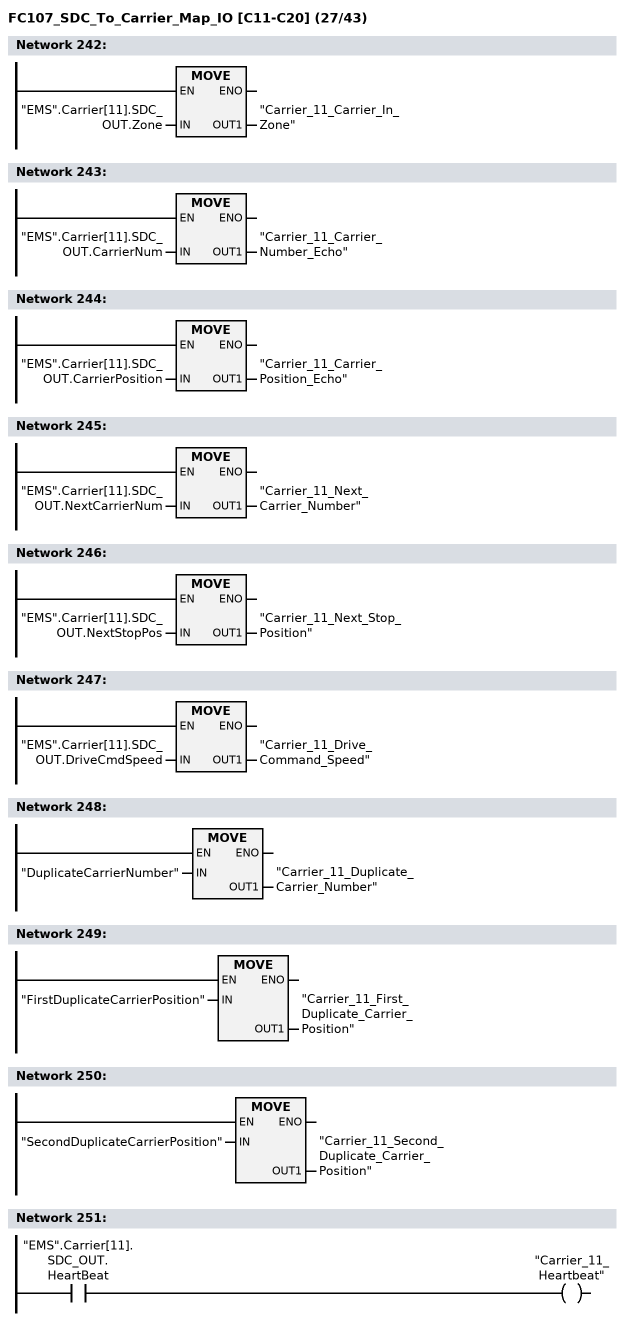
   RUNG wire#powerrail
      Move(in := "EMS".Carrier[11].SDC_OUT.Zone, out1 => "Carrier_11_Carrier_In_Zone")
   END_RUNG
   // the same network as SCL:
   "Carrier_11_Carrier_In_Zone" := "EMS".Carrier[11].SDC_OUT.Zone;
END_REGION

REGION Network 243
   RUNG wire#powerrail
      Move(in := "EMS".Carrier[11].SDC_OUT.CarrierNum, out1 => "Carrier_11_Carrier_Number_Echo")
   END_RUNG
   // the same network as SCL:
   "Carrier_11_Carrier_Number_Echo" := "EMS".Carrier[11].SDC_OUT.CarrierNum;
END_REGION

REGION Network 244
   RUNG wire#powerrail
      Move(in := "EMS".Carrier[11].SDC_OUT.CarrierPosition, out1 => "Carrier_11_Carrier_Position_Echo")
   END_RUNG
   // the same network as SCL:
   "Carrier_11_Carrier_Position_Echo" := "EMS".Carrier[11].SDC_OUT.CarrierPosition;
END_REGION

REGION Network 245
   RUNG wire#powerrail
      Move(in := "EMS".Carrier[11].SDC_OUT.NextCarrierNum, out1 => "Carrier_11_Next_Carrier_Number")
   END_RUNG
   // the same network as SCL:
   "Carrier_11_Next_Carrier_Number" := "EMS".Carrier[11].SDC_OUT.NextCarrierNum;
END_REGION

REGION Network 246
   RUNG wire#powerrail
      Move(in := "EMS".Carrier[11].SDC_OUT.NextStopPos, out1 => "Carrier_11_Next_Stop_Position")
   END_RUNG
   // the same network as SCL:
   "Carrier_11_Next_Stop_Position" := "EMS".Carrier[11].SDC_OUT.NextStopPos;
END_REGION

REGION Network 247
   RUNG wire#powerrail
      Move(in := "EMS".Carrier[11].SDC_OUT.DriveCmdSpeed, out1 => "Carrier_11_Drive_Command_Speed")
   END_RUNG
   // the same network as SCL:
   "Carrier_11_Drive_Command_Speed" := "EMS".Carrier[11].SDC_OUT.DriveCmdSpeed;
END_REGION

REGION Network 248
   RUNG wire#powerrail
      Move(in := "DuplicateCarrierNumber", out1 => "Carrier_11_Duplicate_Carrier_Number")
   END_RUNG
   // the same network as SCL:
   "Carrier_11_Duplicate_Carrier_Number" := "DuplicateCarrierNumber";
END_REGION

REGION Network 249
   RUNG wire#powerrail
      Move(in := "FirstDuplicateCarrierPosition", out1 => "Carrier_11_First_Duplicate_Carrier_Position")
   END_RUNG
   // the same network as SCL:
   "Carrier_11_First_Duplicate_Carrier_Position" := "FirstDuplicateCarrierPosition";
END_REGION

REGION Network 250
   RUNG wire#powerrail
      Move(in := "SecondDuplicateCarrierPosition", out1 => "Carrier_11_Second_Duplicate_Carrier_Position")
   END_RUNG
   // the same network as SCL:
   "Carrier_11_Second_Duplicate_Carrier_Position" := "SecondDuplicateCarrierPosition";
END_REGION

REGION Network 251
   RUNG wire#powerrail
      Contact( "EMS".Carrier[11].SDC_OUT.HeartBeat )
      Coil( "Carrier_11_Heartbeat" )
   END_RUNG
   // the same network as SCL:
   "Carrier_11_Heartbeat" := "EMS".Carrier[11].SDC_OUT.HeartBeat;
END_REGION

REGION Network 252
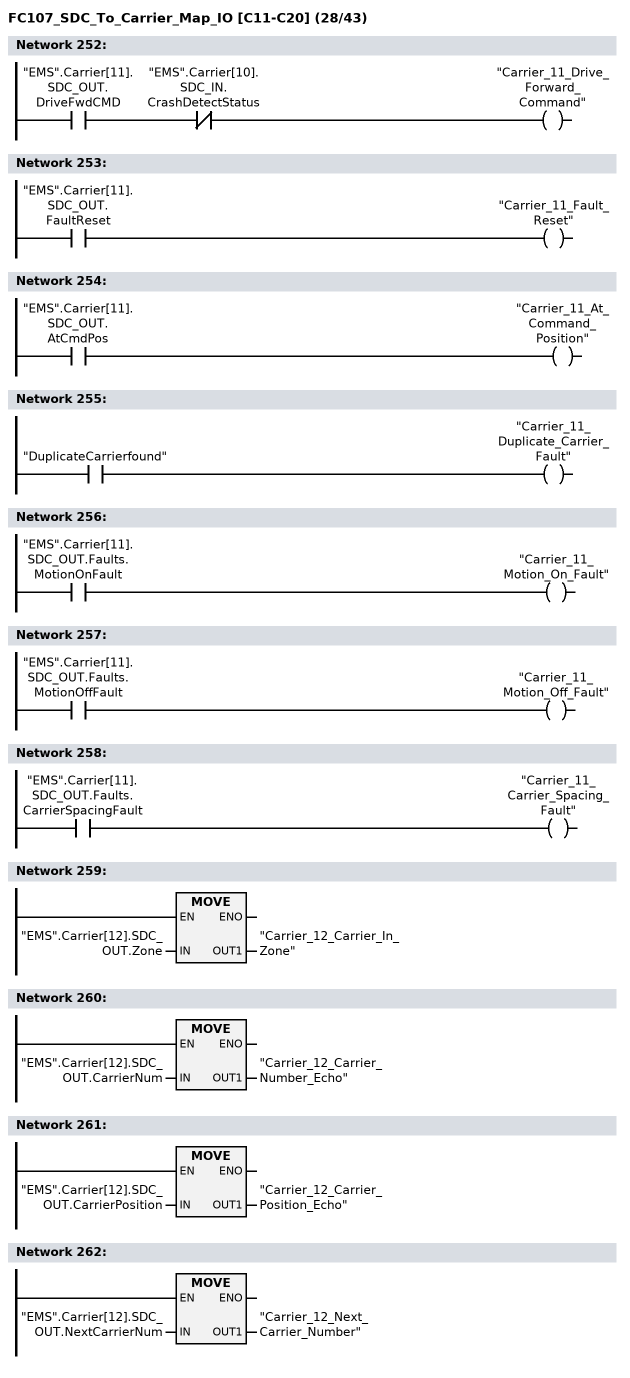
   RUNG wire#powerrail
      Contact( "EMS".Carrier[11].SDC_OUT.DriveFwdCMD )
      I_Contact( "EMS".Carrier[10].SDC_IN.CrashDetectStatus )
      Coil( "Carrier_11_Drive_Forward_Command" )
   END_RUNG
   // the same network as SCL:
   "Carrier_11_Drive_Forward_Command" := "EMS".Carrier[11].SDC_OUT.DriveFwdCMD AND NOT "EMS".Carrier[10].SDC_IN.CrashDetectStatus;
END_REGION

REGION Network 253
   RUNG wire#powerrail
      Contact( "EMS".Carrier[11].SDC_OUT.FaultReset )
      Coil( "Carrier_11_Fault_Reset" )
   END_RUNG
   // the same network as SCL:
   "Carrier_11_Fault_Reset" := "EMS".Carrier[11].SDC_OUT.FaultReset;
END_REGION

REGION Network 254
   RUNG wire#powerrail
      Contact( "EMS".Carrier[11].SDC_OUT.AtCmdPos )
      Coil( "Carrier_11_At_Command_Position" )
   END_RUNG
   // the same network as SCL:
   "Carrier_11_At_Command_Position" := "EMS".Carrier[11].SDC_OUT.AtCmdPos;
END_REGION

REGION Network 255
   RUNG wire#powerrail
      Contact( "DuplicateCarrierfound" )
      Coil( "Carrier_11_Duplicate_Carrier_Fault" )
   END_RUNG
   // the same network as SCL:
   "Carrier_11_Duplicate_Carrier_Fault" := "DuplicateCarrierfound";
END_REGION

REGION Network 256
   RUNG wire#powerrail
      Contact( "EMS".Carrier[11].SDC_OUT.Faults.MotionOnFault )
      Coil( "Carrier_11_Motion_On_Fault" )
   END_RUNG
   // the same network as SCL:
   "Carrier_11_Motion_On_Fault" := "EMS".Carrier[11].SDC_OUT.Faults.MotionOnFault;
END_REGION

REGION Network 257
   RUNG wire#powerrail
      Contact( "EMS".Carrier[11].SDC_OUT.Faults.MotionOffFault )
      Coil( "Carrier_11_Motion_Off_Fault" )
   END_RUNG
   // the same network as SCL:
   "Carrier_11_Motion_Off_Fault" := "EMS".Carrier[11].SDC_OUT.Faults.MotionOffFault;
END_REGION

REGION Network 258
   RUNG wire#powerrail
      Contact( "EMS".Carrier[11].SDC_OUT.Faults.CarrierSpacingFault )
      Coil( "Carrier_11_Carrier_Spacing_Fault" )
   END_RUNG
   // the same network as SCL:
   "Carrier_11_Carrier_Spacing_Fault" := "EMS".Carrier[11].SDC_OUT.Faults.CarrierSpacingFault;
END_REGION

REGION Network 259
   RUNG wire#powerrail
      Move(in := "EMS".Carrier[12].SDC_OUT.Zone, out1 => "Carrier_12_Carrier_In_Zone")
   END_RUNG
   // the same network as SCL:
   "Carrier_12_Carrier_In_Zone" := "EMS".Carrier[12].SDC_OUT.Zone;
END_REGION

REGION Network 260
   RUNG wire#powerrail
      Move(in := "EMS".Carrier[12].SDC_OUT.CarrierNum, out1 => "Carrier_12_Carrier_Number_Echo")
   END_RUNG
   // the same network as SCL:
   "Carrier_12_Carrier_Number_Echo" := "EMS".Carrier[12].SDC_OUT.CarrierNum;
END_REGION

REGION Network 261
   RUNG wire#powerrail
      Move(in := "EMS".Carrier[12].SDC_OUT.CarrierPosition, out1 => "Carrier_12_Carrier_Position_Echo")
   END_RUNG
   // the same network as SCL:
   "Carrier_12_Carrier_Position_Echo" := "EMS".Carrier[12].SDC_OUT.CarrierPosition;
END_REGION

REGION Network 262
   RUNG wire#powerrail
      Move(in := "EMS".Carrier[12].SDC_OUT.NextCarrierNum, out1 => "Carrier_12_Next_Carrier_Number")
   END_RUNG
   // the same network as SCL:
   "Carrier_12_Next_Carrier_Number" := "EMS".Carrier[12].SDC_OUT.NextCarrierNum;
END_REGION

REGION Network 263
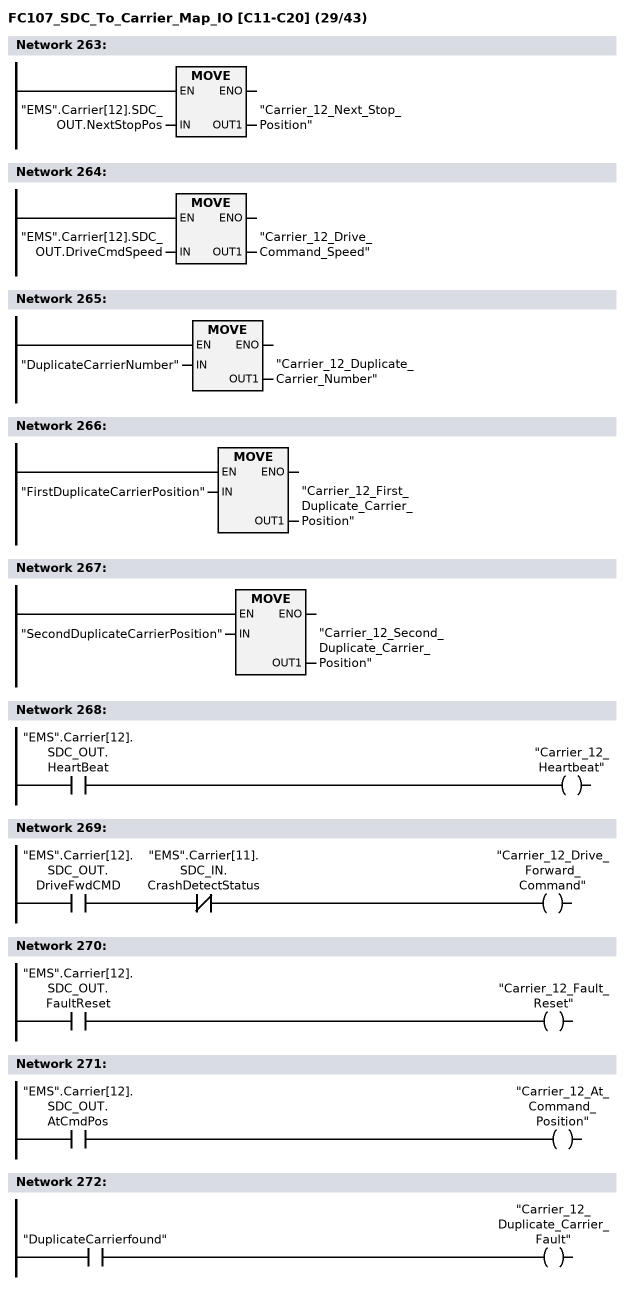
   RUNG wire#powerrail
      Move(in := "EMS".Carrier[12].SDC_OUT.NextStopPos, out1 => "Carrier_12_Next_Stop_Position")
   END_RUNG
   // the same network as SCL:
   "Carrier_12_Next_Stop_Position" := "EMS".Carrier[12].SDC_OUT.NextStopPos;
END_REGION

REGION Network 264
   RUNG wire#powerrail
      Move(in := "EMS".Carrier[12].SDC_OUT.DriveCmdSpeed, out1 => "Carrier_12_Drive_Command_Speed")
   END_RUNG
   // the same network as SCL:
   "Carrier_12_Drive_Command_Speed" := "EMS".Carrier[12].SDC_OUT.DriveCmdSpeed;
END_REGION

REGION Network 265
   RUNG wire#powerrail
      Move(in := "DuplicateCarrierNumber", out1 => "Carrier_12_Duplicate_Carrier_Number")
   END_RUNG
   // the same network as SCL:
   "Carrier_12_Duplicate_Carrier_Number" := "DuplicateCarrierNumber";
END_REGION

REGION Network 266
   RUNG wire#powerrail
      Move(in := "FirstDuplicateCarrierPosition", out1 => "Carrier_12_First_Duplicate_Carrier_Position")
   END_RUNG
   // the same network as SCL:
   "Carrier_12_First_Duplicate_Carrier_Position" := "FirstDuplicateCarrierPosition";
END_REGION

REGION Network 267
   RUNG wire#powerrail
      Move(in := "SecondDuplicateCarrierPosition", out1 => "Carrier_12_Second_Duplicate_Carrier_Position")
   END_RUNG
   // the same network as SCL:
   "Carrier_12_Second_Duplicate_Carrier_Position" := "SecondDuplicateCarrierPosition";
END_REGION

REGION Network 268
   RUNG wire#powerrail
      Contact( "EMS".Carrier[12].SDC_OUT.HeartBeat )
      Coil( "Carrier_12_Heartbeat" )
   END_RUNG
   // the same network as SCL:
   "Carrier_12_Heartbeat" := "EMS".Carrier[12].SDC_OUT.HeartBeat;
END_REGION

REGION Network 269
   RUNG wire#powerrail
      Contact( "EMS".Carrier[12].SDC_OUT.DriveFwdCMD )
      I_Contact( "EMS".Carrier[11].SDC_IN.CrashDetectStatus )
      Coil( "Carrier_12_Drive_Forward_Command" )
   END_RUNG
   // the same network as SCL:
   "Carrier_12_Drive_Forward_Command" := "EMS".Carrier[12].SDC_OUT.DriveFwdCMD AND NOT "EMS".Carrier[11].SDC_IN.CrashDetectStatus;
END_REGION

REGION Network 270
   RUNG wire#powerrail
      Contact( "EMS".Carrier[12].SDC_OUT.FaultReset )
      Coil( "Carrier_12_Fault_Reset" )
   END_RUNG
   // the same network as SCL:
   "Carrier_12_Fault_Reset" := "EMS".Carrier[12].SDC_OUT.FaultReset;
END_REGION

REGION Network 271
   RUNG wire#powerrail
      Contact( "EMS".Carrier[12].SDC_OUT.AtCmdPos )
      Coil( "Carrier_12_At_Command_Position" )
   END_RUNG
   // the same network as SCL:
   "Carrier_12_At_Command_Position" := "EMS".Carrier[12].SDC_OUT.AtCmdPos;
END_REGION

REGION Network 272
   RUNG wire#powerrail
      Contact( "DuplicateCarrierfound" )
      Coil( "Carrier_12_Duplicate_Carrier_Fault" )
   END_RUNG
   // the same network as SCL:
   "Carrier_12_Duplicate_Carrier_Fault" := "DuplicateCarrierfound";
END_REGION

REGION Network 273
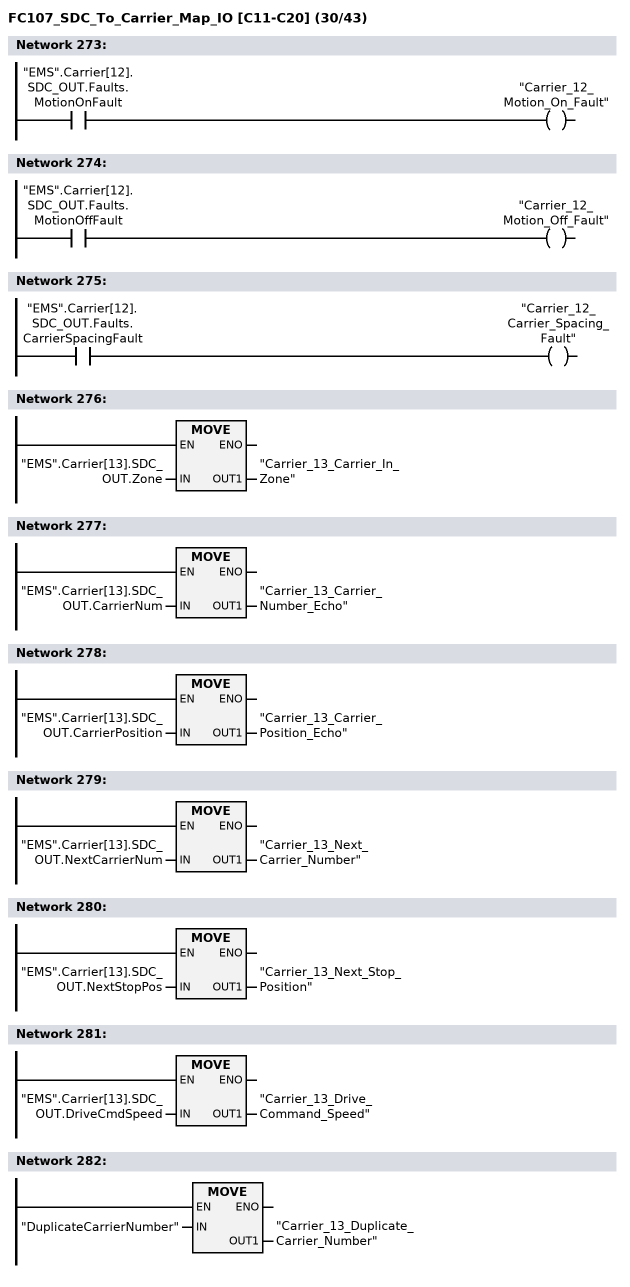
   RUNG wire#powerrail
      Contact( "EMS".Carrier[12].SDC_OUT.Faults.MotionOnFault )
      Coil( "Carrier_12_Motion_On_Fault" )
   END_RUNG
   // the same network as SCL:
   "Carrier_12_Motion_On_Fault" := "EMS".Carrier[12].SDC_OUT.Faults.MotionOnFault;
END_REGION

REGION Network 274
   RUNG wire#powerrail
      Contact( "EMS".Carrier[12].SDC_OUT.Faults.MotionOffFault )
      Coil( "Carrier_12_Motion_Off_Fault" )
   END_RUNG
   // the same network as SCL:
   "Carrier_12_Motion_Off_Fault" := "EMS".Carrier[12].SDC_OUT.Faults.MotionOffFault;
END_REGION

REGION Network 275
   RUNG wire#powerrail
      Contact( "EMS".Carrier[12].SDC_OUT.Faults.CarrierSpacingFault )
      Coil( "Carrier_12_Carrier_Spacing_Fault" )
   END_RUNG
   // the same network as SCL:
   "Carrier_12_Carrier_Spacing_Fault" := "EMS".Carrier[12].SDC_OUT.Faults.CarrierSpacingFault;
END_REGION

REGION Network 276
   RUNG wire#powerrail
      Move(in := "EMS".Carrier[13].SDC_OUT.Zone, out1 => "Carrier_13_Carrier_In_Zone")
   END_RUNG
   // the same network as SCL:
   "Carrier_13_Carrier_In_Zone" := "EMS".Carrier[13].SDC_OUT.Zone;
END_REGION

REGION Network 277
   RUNG wire#powerrail
      Move(in := "EMS".Carrier[13].SDC_OUT.CarrierNum, out1 => "Carrier_13_Carrier_Number_Echo")
   END_RUNG
   // the same network as SCL:
   "Carrier_13_Carrier_Number_Echo" := "EMS".Carrier[13].SDC_OUT.CarrierNum;
END_REGION

REGION Network 278
   RUNG wire#powerrail
      Move(in := "EMS".Carrier[13].SDC_OUT.CarrierPosition, out1 => "Carrier_13_Carrier_Position_Echo")
   END_RUNG
   // the same network as SCL:
   "Carrier_13_Carrier_Position_Echo" := "EMS".Carrier[13].SDC_OUT.CarrierPosition;
END_REGION

REGION Network 279
   RUNG wire#powerrail
      Move(in := "EMS".Carrier[13].SDC_OUT.NextCarrierNum, out1 => "Carrier_13_Next_Carrier_Number")
   END_RUNG
   // the same network as SCL:
   "Carrier_13_Next_Carrier_Number" := "EMS".Carrier[13].SDC_OUT.NextCarrierNum;
END_REGION

REGION Network 280
   RUNG wire#powerrail
      Move(in := "EMS".Carrier[13].SDC_OUT.NextStopPos, out1 => "Carrier_13_Next_Stop_Position")
   END_RUNG
   // the same network as SCL:
   "Carrier_13_Next_Stop_Position" := "EMS".Carrier[13].SDC_OUT.NextStopPos;
END_REGION

REGION Network 281
   RUNG wire#powerrail
      Move(in := "EMS".Carrier[13].SDC_OUT.DriveCmdSpeed, out1 => "Carrier_13_Drive_Command_Speed")
   END_RUNG
   // the same network as SCL:
   "Carrier_13_Drive_Command_Speed" := "EMS".Carrier[13].SDC_OUT.DriveCmdSpeed;
END_REGION

REGION Network 282
   RUNG wire#powerrail
      Move(in := "DuplicateCarrierNumber", out1 => "Carrier_13_Duplicate_Carrier_Number")
   END_RUNG
   // the same network as SCL:
   "Carrier_13_Duplicate_Carrier_Number" := "DuplicateCarrierNumber";
END_REGION

REGION Network 283
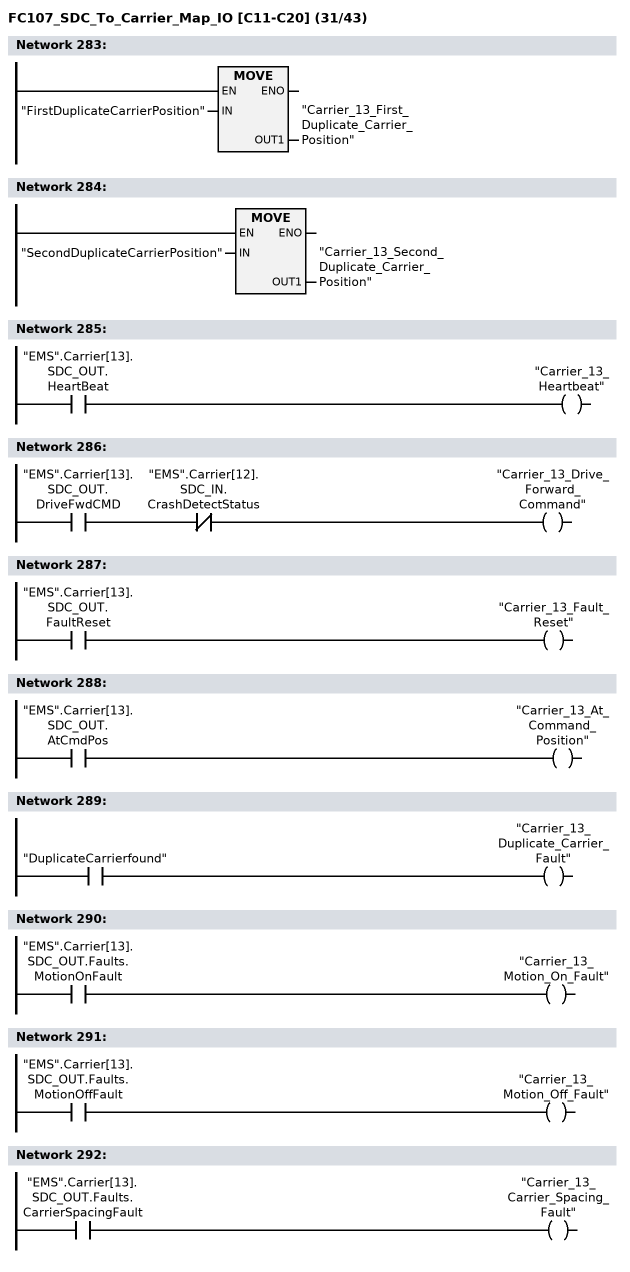
   RUNG wire#powerrail
      Move(in := "FirstDuplicateCarrierPosition", out1 => "Carrier_13_First_Duplicate_Carrier_Position")
   END_RUNG
   // the same network as SCL:
   "Carrier_13_First_Duplicate_Carrier_Position" := "FirstDuplicateCarrierPosition";
END_REGION

REGION Network 284
   RUNG wire#powerrail
      Move(in := "SecondDuplicateCarrierPosition", out1 => "Carrier_13_Second_Duplicate_Carrier_Position")
   END_RUNG
   // the same network as SCL:
   "Carrier_13_Second_Duplicate_Carrier_Position" := "SecondDuplicateCarrierPosition";
END_REGION

REGION Network 285
   RUNG wire#powerrail
      Contact( "EMS".Carrier[13].SDC_OUT.HeartBeat )
      Coil( "Carrier_13_Heartbeat" )
   END_RUNG
   // the same network as SCL:
   "Carrier_13_Heartbeat" := "EMS".Carrier[13].SDC_OUT.HeartBeat;
END_REGION

REGION Network 286
   RUNG wire#powerrail
      Contact( "EMS".Carrier[13].SDC_OUT.DriveFwdCMD )
      I_Contact( "EMS".Carrier[12].SDC_IN.CrashDetectStatus )
      Coil( "Carrier_13_Drive_Forward_Command" )
   END_RUNG
   // the same network as SCL:
   "Carrier_13_Drive_Forward_Command" := "EMS".Carrier[13].SDC_OUT.DriveFwdCMD AND NOT "EMS".Carrier[12].SDC_IN.CrashDetectStatus;
END_REGION

REGION Network 287
   RUNG wire#powerrail
      Contact( "EMS".Carrier[13].SDC_OUT.FaultReset )
      Coil( "Carrier_13_Fault_Reset" )
   END_RUNG
   // the same network as SCL:
   "Carrier_13_Fault_Reset" := "EMS".Carrier[13].SDC_OUT.FaultReset;
END_REGION

REGION Network 288
   RUNG wire#powerrail
      Contact( "EMS".Carrier[13].SDC_OUT.AtCmdPos )
      Coil( "Carrier_13_At_Command_Position" )
   END_RUNG
   // the same network as SCL:
   "Carrier_13_At_Command_Position" := "EMS".Carrier[13].SDC_OUT.AtCmdPos;
END_REGION

REGION Network 289
   RUNG wire#powerrail
      Contact( "DuplicateCarrierfound" )
      Coil( "Carrier_13_Duplicate_Carrier_Fault" )
   END_RUNG
   // the same network as SCL:
   "Carrier_13_Duplicate_Carrier_Fault" := "DuplicateCarrierfound";
END_REGION

REGION Network 290
   RUNG wire#powerrail
      Contact( "EMS".Carrier[13].SDC_OUT.Faults.MotionOnFault )
      Coil( "Carrier_13_Motion_On_Fault" )
   END_RUNG
   // the same network as SCL:
   "Carrier_13_Motion_On_Fault" := "EMS".Carrier[13].SDC_OUT.Faults.MotionOnFault;
END_REGION

REGION Network 291
   RUNG wire#powerrail
      Contact( "EMS".Carrier[13].SDC_OUT.Faults.MotionOffFault )
      Coil( "Carrier_13_Motion_Off_Fault" )
   END_RUNG
   // the same network as SCL:
   "Carrier_13_Motion_Off_Fault" := "EMS".Carrier[13].SDC_OUT.Faults.MotionOffFault;
END_REGION

REGION Network 292
   RUNG wire#powerrail
      Contact( "EMS".Carrier[13].SDC_OUT.Faults.CarrierSpacingFault )
      Coil( "Carrier_13_Carrier_Spacing_Fault" )
   END_RUNG
   // the same network as SCL:
   "Carrier_13_Carrier_Spacing_Fault" := "EMS".Carrier[13].SDC_OUT.Faults.CarrierSpacingFault;
END_REGION

REGION Network 293
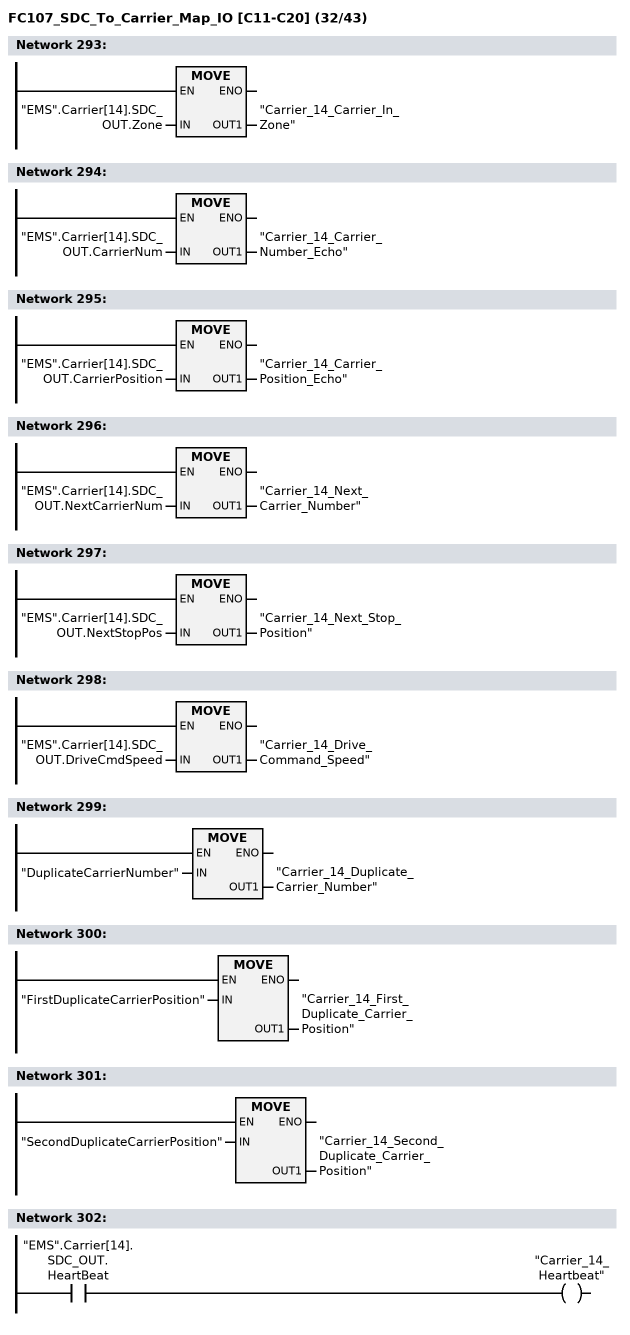
   RUNG wire#powerrail
      Move(in := "EMS".Carrier[14].SDC_OUT.Zone, out1 => "Carrier_14_Carrier_In_Zone")
   END_RUNG
   // the same network as SCL:
   "Carrier_14_Carrier_In_Zone" := "EMS".Carrier[14].SDC_OUT.Zone;
END_REGION

REGION Network 294
   RUNG wire#powerrail
      Move(in := "EMS".Carrier[14].SDC_OUT.CarrierNum, out1 => "Carrier_14_Carrier_Number_Echo")
   END_RUNG
   // the same network as SCL:
   "Carrier_14_Carrier_Number_Echo" := "EMS".Carrier[14].SDC_OUT.CarrierNum;
END_REGION

REGION Network 295
   RUNG wire#powerrail
      Move(in := "EMS".Carrier[14].SDC_OUT.CarrierPosition, out1 => "Carrier_14_Carrier_Position_Echo")
   END_RUNG
   // the same network as SCL:
   "Carrier_14_Carrier_Position_Echo" := "EMS".Carrier[14].SDC_OUT.CarrierPosition;
END_REGION

REGION Network 296
   RUNG wire#powerrail
      Move(in := "EMS".Carrier[14].SDC_OUT.NextCarrierNum, out1 => "Carrier_14_Next_Carrier_Number")
   END_RUNG
   // the same network as SCL:
   "Carrier_14_Next_Carrier_Number" := "EMS".Carrier[14].SDC_OUT.NextCarrierNum;
END_REGION

REGION Network 297
   RUNG wire#powerrail
      Move(in := "EMS".Carrier[14].SDC_OUT.NextStopPos, out1 => "Carrier_14_Next_Stop_Position")
   END_RUNG
   // the same network as SCL:
   "Carrier_14_Next_Stop_Position" := "EMS".Carrier[14].SDC_OUT.NextStopPos;
END_REGION

REGION Network 298
   RUNG wire#powerrail
      Move(in := "EMS".Carrier[14].SDC_OUT.DriveCmdSpeed, out1 => "Carrier_14_Drive_Command_Speed")
   END_RUNG
   // the same network as SCL:
   "Carrier_14_Drive_Command_Speed" := "EMS".Carrier[14].SDC_OUT.DriveCmdSpeed;
END_REGION

REGION Network 299
   RUNG wire#powerrail
      Move(in := "DuplicateCarrierNumber", out1 => "Carrier_14_Duplicate_Carrier_Number")
   END_RUNG
   // the same network as SCL:
   "Carrier_14_Duplicate_Carrier_Number" := "DuplicateCarrierNumber";
END_REGION

REGION Network 300
   RUNG wire#powerrail
      Move(in := "FirstDuplicateCarrierPosition", out1 => "Carrier_14_First_Duplicate_Carrier_Position")
   END_RUNG
   // the same network as SCL:
   "Carrier_14_First_Duplicate_Carrier_Position" := "FirstDuplicateCarrierPosition";
END_REGION

REGION Network 301
   RUNG wire#powerrail
      Move(in := "SecondDuplicateCarrierPosition", out1 => "Carrier_14_Second_Duplicate_Carrier_Position")
   END_RUNG
   // the same network as SCL:
   "Carrier_14_Second_Duplicate_Carrier_Position" := "SecondDuplicateCarrierPosition";
END_REGION

REGION Network 302
   RUNG wire#powerrail
      Contact( "EMS".Carrier[14].SDC_OUT.HeartBeat )
      Coil( "Carrier_14_Heartbeat" )
   END_RUNG
   // the same network as SCL:
   "Carrier_14_Heartbeat" := "EMS".Carrier[14].SDC_OUT.HeartBeat;
END_REGION

REGION Network 303
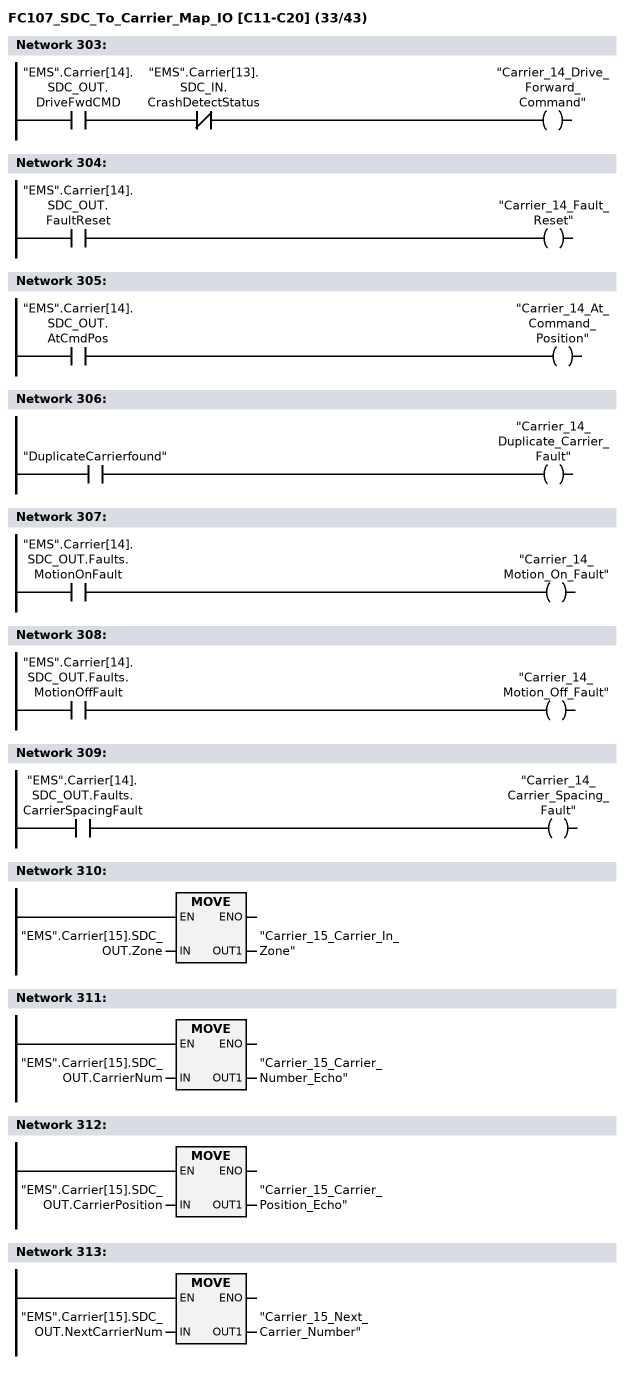
   RUNG wire#powerrail
      Contact( "EMS".Carrier[14].SDC_OUT.DriveFwdCMD )
      I_Contact( "EMS".Carrier[13].SDC_IN.CrashDetectStatus )
      Coil( "Carrier_14_Drive_Forward_Command" )
   END_RUNG
   // the same network as SCL:
   "Carrier_14_Drive_Forward_Command" := "EMS".Carrier[14].SDC_OUT.DriveFwdCMD AND NOT "EMS".Carrier[13].SDC_IN.CrashDetectStatus;
END_REGION

REGION Network 304
   RUNG wire#powerrail
      Contact( "EMS".Carrier[14].SDC_OUT.FaultReset )
      Coil( "Carrier_14_Fault_Reset" )
   END_RUNG
   // the same network as SCL:
   "Carrier_14_Fault_Reset" := "EMS".Carrier[14].SDC_OUT.FaultReset;
END_REGION

REGION Network 305
   RUNG wire#powerrail
      Contact( "EMS".Carrier[14].SDC_OUT.AtCmdPos )
      Coil( "Carrier_14_At_Command_Position" )
   END_RUNG
   // the same network as SCL:
   "Carrier_14_At_Command_Position" := "EMS".Carrier[14].SDC_OUT.AtCmdPos;
END_REGION

REGION Network 306
   RUNG wire#powerrail
      Contact( "DuplicateCarrierfound" )
      Coil( "Carrier_14_Duplicate_Carrier_Fault" )
   END_RUNG
   // the same network as SCL:
   "Carrier_14_Duplicate_Carrier_Fault" := "DuplicateCarrierfound";
END_REGION

REGION Network 307
   RUNG wire#powerrail
      Contact( "EMS".Carrier[14].SDC_OUT.Faults.MotionOnFault )
      Coil( "Carrier_14_Motion_On_Fault" )
   END_RUNG
   // the same network as SCL:
   "Carrier_14_Motion_On_Fault" := "EMS".Carrier[14].SDC_OUT.Faults.MotionOnFault;
END_REGION

REGION Network 308
   RUNG wire#powerrail
      Contact( "EMS".Carrier[14].SDC_OUT.Faults.MotionOffFault )
      Coil( "Carrier_14_Motion_Off_Fault" )
   END_RUNG
   // the same network as SCL:
   "Carrier_14_Motion_Off_Fault" := "EMS".Carrier[14].SDC_OUT.Faults.MotionOffFault;
END_REGION

REGION Network 309
   RUNG wire#powerrail
      Contact( "EMS".Carrier[14].SDC_OUT.Faults.CarrierSpacingFault )
      Coil( "Carrier_14_Carrier_Spacing_Fault" )
   END_RUNG
   // the same network as SCL:
   "Carrier_14_Carrier_Spacing_Fault" := "EMS".Carrier[14].SDC_OUT.Faults.CarrierSpacingFault;
END_REGION

REGION Network 310
   RUNG wire#powerrail
      Move(in := "EMS".Carrier[15].SDC_OUT.Zone, out1 => "Carrier_15_Carrier_In_Zone")
   END_RUNG
   // the same network as SCL:
   "Carrier_15_Carrier_In_Zone" := "EMS".Carrier[15].SDC_OUT.Zone;
END_REGION

REGION Network 311
   RUNG wire#powerrail
      Move(in := "EMS".Carrier[15].SDC_OUT.CarrierNum, out1 => "Carrier_15_Carrier_Number_Echo")
   END_RUNG
   // the same network as SCL:
   "Carrier_15_Carrier_Number_Echo" := "EMS".Carrier[15].SDC_OUT.CarrierNum;
END_REGION

REGION Network 312
   RUNG wire#powerrail
      Move(in := "EMS".Carrier[15].SDC_OUT.CarrierPosition, out1 => "Carrier_15_Carrier_Position_Echo")
   END_RUNG
   // the same network as SCL:
   "Carrier_15_Carrier_Position_Echo" := "EMS".Carrier[15].SDC_OUT.CarrierPosition;
END_REGION

REGION Network 313
   RUNG wire#powerrail
      Move(in := "EMS".Carrier[15].SDC_OUT.NextCarrierNum, out1 => "Carrier_15_Next_Carrier_Number")
   END_RUNG
   // the same network as SCL:
   "Carrier_15_Next_Carrier_Number" := "EMS".Carrier[15].SDC_OUT.NextCarrierNum;
END_REGION

REGION Network 314
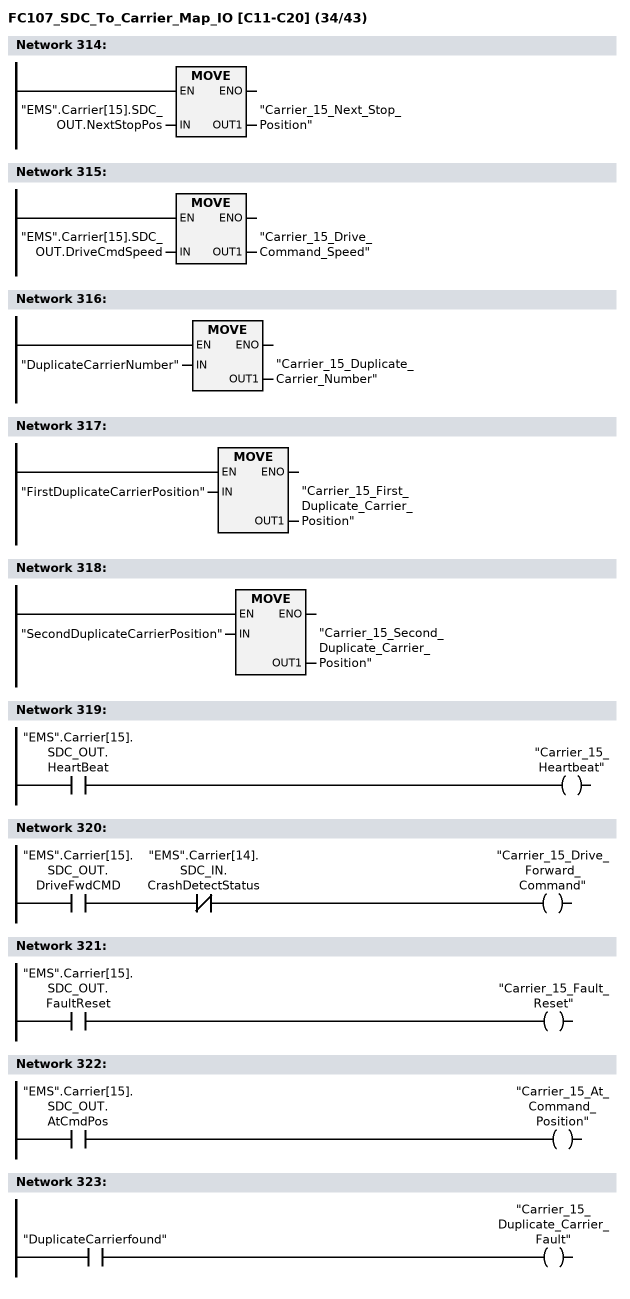
   RUNG wire#powerrail
      Move(in := "EMS".Carrier[15].SDC_OUT.NextStopPos, out1 => "Carrier_15_Next_Stop_Position")
   END_RUNG
   // the same network as SCL:
   "Carrier_15_Next_Stop_Position" := "EMS".Carrier[15].SDC_OUT.NextStopPos;
END_REGION

REGION Network 315
   RUNG wire#powerrail
      Move(in := "EMS".Carrier[15].SDC_OUT.DriveCmdSpeed, out1 => "Carrier_15_Drive_Command_Speed")
   END_RUNG
   // the same network as SCL:
   "Carrier_15_Drive_Command_Speed" := "EMS".Carrier[15].SDC_OUT.DriveCmdSpeed;
END_REGION

REGION Network 316
   RUNG wire#powerrail
      Move(in := "DuplicateCarrierNumber", out1 => "Carrier_15_Duplicate_Carrier_Number")
   END_RUNG
   // the same network as SCL:
   "Carrier_15_Duplicate_Carrier_Number" := "DuplicateCarrierNumber";
END_REGION

REGION Network 317
   RUNG wire#powerrail
      Move(in := "FirstDuplicateCarrierPosition", out1 => "Carrier_15_First_Duplicate_Carrier_Position")
   END_RUNG
   // the same network as SCL:
   "Carrier_15_First_Duplicate_Carrier_Position" := "FirstDuplicateCarrierPosition";
END_REGION

REGION Network 318
   RUNG wire#powerrail
      Move(in := "SecondDuplicateCarrierPosition", out1 => "Carrier_15_Second_Duplicate_Carrier_Position")
   END_RUNG
   // the same network as SCL:
   "Carrier_15_Second_Duplicate_Carrier_Position" := "SecondDuplicateCarrierPosition";
END_REGION

REGION Network 319
   RUNG wire#powerrail
      Contact( "EMS".Carrier[15].SDC_OUT.HeartBeat )
      Coil( "Carrier_15_Heartbeat" )
   END_RUNG
   // the same network as SCL:
   "Carrier_15_Heartbeat" := "EMS".Carrier[15].SDC_OUT.HeartBeat;
END_REGION

REGION Network 320
   RUNG wire#powerrail
      Contact( "EMS".Carrier[15].SDC_OUT.DriveFwdCMD )
      I_Contact( "EMS".Carrier[14].SDC_IN.CrashDetectStatus )
      Coil( "Carrier_15_Drive_Forward_Command" )
   END_RUNG
   // the same network as SCL:
   "Carrier_15_Drive_Forward_Command" := "EMS".Carrier[15].SDC_OUT.DriveFwdCMD AND NOT "EMS".Carrier[14].SDC_IN.CrashDetectStatus;
END_REGION

REGION Network 321
   RUNG wire#powerrail
      Contact( "EMS".Carrier[15].SDC_OUT.FaultReset )
      Coil( "Carrier_15_Fault_Reset" )
   END_RUNG
   // the same network as SCL:
   "Carrier_15_Fault_Reset" := "EMS".Carrier[15].SDC_OUT.FaultReset;
END_REGION

REGION Network 322
   RUNG wire#powerrail
      Contact( "EMS".Carrier[15].SDC_OUT.AtCmdPos )
      Coil( "Carrier_15_At_Command_Position" )
   END_RUNG
   // the same network as SCL:
   "Carrier_15_At_Command_Position" := "EMS".Carrier[15].SDC_OUT.AtCmdPos;
END_REGION

REGION Network 323
   RUNG wire#powerrail
      Contact( "DuplicateCarrierfound" )
      Coil( "Carrier_15_Duplicate_Carrier_Fault" )
   END_RUNG
   // the same network as SCL:
   "Carrier_15_Duplicate_Carrier_Fault" := "DuplicateCarrierfound";
END_REGION

REGION Network 324